(* Logix 5000 project; controller PLC_MCC1201_220AP1 vendor 1 type 14 code 164 rev 35.11; software revision 35.00; part 5 of 25 *)
(* tags used below, declared in another part *)
   B3 : DINT[102];
   B52 : DINT[100];
   GP_OB_InitializeMain : GP_OB_Initialize;
   HMI_Alarm_Reset : BOOL;   // HMI_Alarm_Reset
   HMI_MAN_CMD_WR : UDT_MAN_CMD_WR;
   HOST_DATA_REQ : ALIAS FOR N43[209].0;
   I : INT[128];
   LEHR_SPEED : ALIAS FOR N60[1];
   M202_M1_DR : AXIS_CIP_DRIVE;
   M203_M1_DR : AXIS_CIP_DRIVE;
   M203DROP : MAC_DROPCONV;
   M203DROP_HMR : MAC_DROPCONV_HMR;
   M204_M1_DR : AXIS_CIP_DRIVE;
   M2xx_CONVEYOR : MAC_CONVEYOR[20];
   M2xx_CONVEYOR_IN_MOTION : MAC_CONVEYOR_IN_MOTION[20];
   M2xx_CONVEYOR_OUT_MOTION : MAC_CONVEYOR_OUT_MOTION[20];
   MS_ACCUM : ALIAS FOR N70[1];
   N : ALIAS FOR N15[80];
   N43 : DINT[240];
   N54 : DINT[501];
   N70 : DINT[3];
   N80 : DINT[16];
   O : INT[128];
   REL_CAP_REQUEST : ALIAS FOR I[17].14;
   S : INT[128];
   Status : INT;   // INT tag to retrieve Status value through GSV created during conversion
   T4 : TIMER[100];
   T57 : TIMER[100];
   TMP_dDirection : DINT;
   TMP_rAcc : REAL;
   TMP_rDec : REAL;
   TMP_rSpeed : REAL;
   TMP_xAlwaysOFF : BOOL;
   TMP_xRun : BOOL;
   W_B3 : DINT[7];

   W_CONV_MSG_N7_0 : MESSAGE;   // IFE1_BTW_CNT
        .EN   // btw_enable
        MessageParameters(ServiceCode := 16#004c, LocalElement := W_N7[10], ...)
   W_CONV_MSG_N7_120 : MESSAGE;   // OFE1_CONTROL
        .EN   // BTW_OFE1_ENABLE
        MessageParameters(ServiceCode := 16#004c, LocalElement := W_N7[140], ...)
   W_CONV_MSG_N7_160 : MESSAGE;   // OFE1_BTR_CONTRO
        .EN   // OFE1_BTR_ENABLE
        MessageParameters(ServiceCode := 16#004b, LocalElement := W_N7[180], ...)
   W_CONV_MSG_N7_200 : MESSAGE;   // OFE2_CONTROL
        .EN   // OFE2_BTW_ENABLE
        MessageParameters(ServiceCode := 16#004c, LocalElement := W_N7[220], ...)
   W_CONV_MSG_N7_240 : MESSAGE;   // OFE2_BTR_CONTRO
        .EN   // OFE2_BTR_ENABLE
        MessageParameters(ServiceCode := 16#004b, LocalElement := W_N7[260], ...)
   W_CONV_MSG_N7_280 : MESSAGE;   // OFE3_CONTROL
        .EN   // OFE3_BTW_ENABLE
        MessageParameters(ServiceCode := 16#004c, LocalElement := W_N7[300], ...)
   W_CONV_MSG_N7_32 : MESSAGE;   // IFE1_BTR
        .EN   // BTR_IFE1_ENABLE
        MessageParameters(ServiceCode := 16#004b, LocalElement := W_N7[42], ...)
   W_CONV_MSG_N7_320 : MESSAGE;   // OFE3_BTR_CONTRL
        .EN   // OFE3_BTR_ENABLE
        MessageParameters(ServiceCode := 16#004b, LocalElement := W_N7[340], ...)
   W_CONV_MSG_N7_360 : MESSAGE;   // OFE4_CONTROL
        .EN   // OFE4_BTW_CONTRL
        MessageParameters(ServiceCode := 16#004c, LocalElement := W_N7[380], ...)
   W_CONV_MSG_N7_400 : MESSAGE;   // OFE4_BTR_CONTRL
        .EN   // OFE4_BTR_ENABLE
        MessageParameters(ServiceCode := 16#004b, LocalElement := W_N7[420], ...)
   W_CONV_MSG_N7_60 : MESSAGE;   // IFE2_CONTROL
        .EN   // IFE2_BTW_ENABLE
        MessageParameters(ServiceCode := 16#004c, LocalElement := W_N7[70], ...)
   W_CONV_MSG_N7_92 : MESSAGE;   // IFE2_BTR
        .EN   // BTR_IFE2_ENABLE
        MessageParameters(ServiceCode := 16#004b, LocalElement := W_N7[102], ...)
   W_CONV_PID_N7_440 : PID := (CTL := 1115722368, CT := 1, CA := 1, PE := 1, INI := 1, OLH := 1, DVPA := 1, PVHA := 1, SP := 2048.0, KP := 500.0, BIAS := 2973.0, MAXS := 4095.0, SO := 100.0, MAXO := 100.0, UPD := 1.0, PV := 4095.0, ERR := 2047.0, OUT := 100.0, MAXI := 4095.0, MAXTIE := 4095.0, DATA[1] := 1600.0, DATA[2] := 4095.0, DATA[3] := 2047.0, DATA[4] := 2048.0, DATA[5] := 0.024420025, DATA[6] := 1.0, DATA[7] := 16.0, DATA[8] := 500.0, DATA[11] := 500.0, DATA[16] := 0.024420025);   // Receiving Tank Level Control
   W_CONV_PID_N7_470 : PID := (CTL := 1082168192, CT := 1, PE := 1, INI := 1, OLH := 1, DVPA := 1, PVLA := 1, PVHA := 1, SP := 1845.0, KP := 150.0, KI := 300.0, BIAS := 2045.0, MAXS := 4095.0, SO := 100.0, MAXO := 100.0, UPD := 1.0, ERR := 1845.0, OUT := 100.0, MAXI := 4095.0, MAXTIE := 4095.0, DATA[3] := 1845.0, DATA[4] := 1845.0, DATA[5] := 0.024420025, DATA[6] := 1.0, DATA[7] := 16.0, DATA[8] := 150.0, DATA[9] := 300.0, DATA[11] := 150.0, DATA[12] := 0.008333334, DATA[16] := 0.024420025);   // Washer Water Pressure Cntrl Valve Position
   W_CONV_PID_N7_500 : PID := (CTL := 1082168192, CT := 1, PE := 1, INI := 1, OLH := 1, DVPA := 1, PVLA := 1, PVHA := 1, SP := 2050.0, KP := 250.0, BIAS := 2045.0, MAXS := 4095.0, SO := 100.0, MAXO := 100.0, UPD := 1.0, ERR := 2050.0, OUT := 100.0, MAXI := 4095.0, MAXTIE := 4095.0, DATA[3] := 2050.0, DATA[4] := 2050.0, DATA[5] := 0.024420025, DATA[6] := 1.0, DATA[7] := 16.0, DATA[8] := 250.0, DATA[11] := 250.0, DATA[16] := 0.024420025);   // Dryer Room Airflow (CB2) Fan Actuator Control
   W_CONV_PID_N7_530 : PID := (CTL := 8430720, PE := 1, INI := 1, OLL := 1, DVNA := 1, PVHA := 1, SP := 2073.0, KP := 100.0, KI := 300.0, BIAS := 2047.0, MAXS := 4095.0, MAXO := 100.0, UPD := 1.0, PV := 4095.0, ERR := -2022.0, MAXI := 4095.0, MAXTIE := 4095.0, DATA[1] := -1600.0, DATA[2] := 4095.0, DATA[3] := -2022.0, DATA[4] := 2073.0, DATA[5] := 0.024420025, DATA[6] := 1.0, DATA[7] := 16.0, DATA[8] := 100.0, DATA[9] := 300.0, DATA[11] := 100.0, DATA[12] := 0.0055555557, DATA[16] := 0.024420025);   // Blower CB1 Static Pressure Fan Actuator Control
   W_CONV_PID_N7_560 : PID := (CTL := 8430720, PE := 1, INI := 1, OLL := 1, DVNA := 1, PVHA := 1, SP := 1023.0, KP := 300.0, KI := 300.0, BIAS := 2047.0, MAXS := 4095.0, MAXO := 100.0, UPD := 1.0, PV := 1339.0, ERR := -316.0, MAXI := 4095.0, MAXTIE := 4095.0, DATA[1] := -523.1746, DATA[2] := 1339.0, DATA[3] := -316.0, DATA[4] := 1023.0, DATA[5] := 0.024420025, DATA[6] := 1.0, DATA[7] := 16.0, DATA[8] := 300.0, DATA[9] := 300.0, DATA[11] := 300.0, DATA[12] := 0.016666668, DATA[16] := 0.024420025);   // RO Heating Coil Temp. Control (HC1)
   W_CONV_PID_N7_590 : PID := (CTL := 1082167936, CT := 1, PE := 1, INI := 1, OLH := 1, DVPA := 1, PVHA := 1, SP := 2559.0, KP := 250.0, KI := 300.0, BIAS := 2047.0, MAXS := 4095.0, SO := 100.0, MAXO := 100.0, UPD := 1.0, PV := 525.0, ERR := 2034.0, OUT := 100.0, MAXI := 4095.0, MAXTIE := 4095.0, DATA[1] := -205.1282, DATA[2] := 525.0, DATA[3] := 2034.0, DATA[4] := 2559.0, DATA[5] := 0.024420025, DATA[6] := 1.0, DATA[7] := 16.0, DATA[8] := 250.0, DATA[9] := 300.0, DATA[11] := 250.0, DATA[12] := 0.013888889, DATA[16] := 0.024420025);   // Eclipse Heating Coil Temp. Control
   W_CONV_PID_N7_620 : PID := (CTL := 1082168192, CT := 1, PE := 1, INI := 1, OLH := 1, DVPA := 1, PVLA := 1, PVHA := 1, SP := 615.0, KP := 500.0, KI := 300.0, BIAS := 2047.0, MAXS := 4095.0, SO := 100.0, MAXO := 100.0, UPD := 1.0, ERR := 615.0, OUT := 100.0, MAXI := 4095.0, MAXTIE := 4095.0, DATA[3] := 615.0, DATA[4] := 615.0, DATA[5] := 0.024420025, DATA[6] := 1.0, DATA[7] := 16.0, DATA[8] := 500.0, DATA[9] := 300.0, DATA[11] := 500.0, DATA[12] := 0.027777778, DATA[16] := 0.024420025);   // Return Water Flow Control Valve Position
   W_CONV_PID_N7_650 : PID := (CTL := 41985152, CA := 1, PE := 1, INI := 1, OLL := 1, DVNA := 1, PVHA := 1, SP := 1971.0, KP := 400.0, KI := 100.0, BIAS := 2047.0, MAXS := 4095.0, MAXO := 100.0, UPD := 1.0, PV := 1713.0, ERR := -258.0, MAXI := 4095.0, MAXTIE := 4095.0, DATA[1] := 669.304, DATA[2] := 1713.0, DATA[3] := -258.0, DATA[4] := 1971.0, DATA[5] := 0.024420025, DATA[6] := 1.0, DATA[7] := 16.0, DATA[8] := 400.0, DATA[9] := 100.0, DATA[11] := 400.0, DATA[12] := 0.06666667, DATA[16] := 0.024420025);   // RO Unit Water Temperature Control
   W_CONV_PID_N7_680 : PID := (CTL := 1082167936, CT := 1, PE := 1, INI := 1, OLH := 1, DVPA := 1, PVHA := 1, SP := 2047.0, KP := 300.0, KI := 300.0, BIAS := 2047.0, MAXS := 4095.0, SO := 100.0, MAXO := 100.0, UPD := 1.0, PV := 439.0, ERR := 1608.0, OUT := 100.0, MAXI := 4095.0, MAXTIE := 4095.0, DATA[1] := -171.52626, DATA[2] := 439.0, DATA[3] := 1608.0, DATA[4] := 2047.0, DATA[5] := 0.024420025, DATA[6] := 1.0, DATA[7] := 16.0, DATA[8] := 300.0, DATA[9] := 300.0, DATA[11] := 300.0, DATA[12] := 0.016666668, DATA[16] := 0.024420025);   // Boiler Water Temperature Control
   W_CONV_PID_N7_710 : PID := (CTL := 1082167936, CT := 1, PE := 1, INI := 1, OLH := 1, DVPA := 1, PVHA := 1, SP := 2047.0, KP := 300.0, KI := 200.0, BIAS := 2047.0, MAXS := 4095.0, SO := 100.0, MAXO := 100.0, UPD := 1.0, PV := 1029.0, ERR := 1018.0, OUT := 100.0, MAXI := 4095.0, MAXTIE := 4095.0, DATA[1] := -402.0513, DATA[2] := 1029.0, DATA[3] := 1018.0, DATA[4] := 2047.0, DATA[5] := 0.024420025, DATA[6] := 1.0, DATA[7] := 16.0, DATA[8] := 300.0, DATA[9] := 200.0, DATA[11] := 300.0, DATA[12] := 0.025, DATA[16] := 0.024420025);   // Mixed Air Control Damper Positioning
   W_CONV_PID_N7_740 : PID := (CTL := 1082168192, CT := 1, PE := 1, INI := 1, OLH := 1, DVPA := 1, PVLA := 1, PVHA := 1, SP := 1024.0, KP := 300.0, KI := 300.0, BIAS := 2047.0, MAXS := 4095.0, SO := 100.0, MAXO := 100.0, UPD := 1.0, ERR := 1024.0, OUT := 100.0, MAXI := 4095.0, MAXTIE := 4095.0, DATA[3] := 1024.0, DATA[4] := 1024.0, DATA[5] := 0.024420025, DATA[6] := 1.0, DATA[7] := 16.0, DATA[8] := 300.0, DATA[9] := 300.0, DATA[11] := 300.0, DATA[12] := 0.016666668, DATA[16] := 0.024420025);   // Dryer Room Temperature Control
   W_CP1_ENABLE : ALIAS FOR W_B3[0].5;
   W_CP1A_START : ALIAS FOR W_O[10].5;
   W_CP1A_STATUS : ALIAS FOR W_I[8].7;
   W_CP1B_START : ALIAS FOR W_O[10].7;
   W_CP1B_STATUS : ALIAS FOR W_I[8].6;
   W_CP2A_START : ALIAS FOR W_O[10].9;
   W_CP2A_STAT : ALIAS FOR W_I[8].4;
   W_CP2B_START : ALIAS FOR W_O[10].11;
   W_CP2B_STAT : ALIAS FOR W_I[8].3;
   W_DRV_OUTPUT : ALIAS FOR W_N7[380];
   W_DRV_PID : ALIAS FOR W_N7[440];
   W_DRYER_AIR_FLOW : ALIAS FOR W_N7[108];
   W_DRYER_PID_OUT : ALIAS FOR W_N7[925];
   W_DRYER_TEMP_PID : ALIAS FOR W_N7[740];
   W_DRYER_TEMP_TMR : ALIAS FOR W_T4[16];
   W_EMER_STOP : ALIAS FOR W_I[8].13;
   W_EMER_STOP_LIGHT : ALIAS FOR W_O[10].10;
   W_F8 : REAL[1];
   W_FAN_CB1_TIMER : ALIAS FOR W_T4[4];
   W_FAN_CB2_TIMER : ALIAS FOR W_T4[5];
   W_FLOW_ENABLE : ALIAS FOR W_B3[0].9;
   W_HC1_SENSOR : ALIAS FOR W_N7[44];
   W_HEATING_AIR_ST : ALIAS FOR W_N7[107];
   W_HX1_BCD_OUT : ALIAS FOR W_N7[917];
   W_HX2_SENSOR : ALIAS FOR W_N7[47];
   W_I : INT[32] := ([8] := 2#0001_0000_0000_0110, [17] := 2#0000_0000_0101_0000);
        [16].8   // ?????????????? RO System Emergency Low Level Photoeye ??????????????
        [16].0   // Pump CP1A Drive Fault
        [16].1   // Pump CP1B Drive Fault
        [16].2   // RO Water Low Feed Pressure
        [16].3   // Reverse Osmosis Pump Motor Auxillary
        [16].4   // Eclipse On Selector at NSG Washer Panel (North)
        [16].5   // Eclipse Off Selector at NSG Washer Panel (North)
        [16].6   // Elipse On Selector at NSG Washer Panel (South)
        [16].7   // Eclipse Off Selector at NSG Washer Panel (South)
        [8].0   // Logical Shutdown Pushbutton
        [8].1   // Process Water Tank Low Level Limit Switch (Honeywell)
        [8].10   // APC Tank Fill Switch
        [8].11   // CB2 Blower Starter Auxillary
        [8].12   // CB1 Blower Starter Auxillary
        [8].13   // RO System Emergency Stop
        [8].14   // Pump CP1 Lead/Lag Switch
        [8].15   // Pump CP2 Lead/Lag Switch
        [8].2   // Process Water Tank High Limit
        [8].3   // CP2B Motor Starter Auxillary Status
        [8].4   // CP2A Motor Starter Auxillary Status
        [8].6   // CP1B Motor Auxillary Status
        [8].7   // CP1A Motor Auxillary Status
        [8].8   // PS1_Switch Pressure Switch
        [8].9   // Recieving Tank Level Switch (Cullet Tunnel)
        [8]   // WASHER INPUTS
        [16]   // WASHER INPUTS
   W_IFE1_BTW_CNT : ALIAS FOR W_N7[0];
   W_IFE1_BTW_DATA : ALIAS FOR W_N7[10];
   W_IFE2_BTR : ALIAS FOR W_N7[92];
   W_IFE2_CONTROL : ALIAS FOR W_N7[60];
   W_IFE2_DATA : ALIAS FOR W_N7[70];
   W_INT_FOR_BCD1 : ALIAS FOR W_N7[911];
   W_LEVEL_SENSOR : ALIAS FOR W_N7[109];
   W_LL_CP1 : ALIAS FOR W_I[8].14;
   W_LL_CP1A_T : ALIAS FOR W_T4[2];
   W_LL_CP1B_T : ALIAS FOR W_T4[3];
   W_LL_CP2 : ALIAS FOR W_I[8].15;
   W_LL_CP2A_T : ALIAS FOR W_T4[0];
   W_LL_CP2B_T : ALIAS FOR W_T4[1];
   W_LL_TIMER : ALIAS FOR W_T4[100];
   W_LOG_SHUTDOWN : ALIAS FOR W_I[8].0;
   W_MA_FAN_SENSOR : ALIAS FOR W_N7[50];
   W_MIX_AIR_PID : ALIAS FOR W_N7[710];
   W_N11 : DINT[10] := ([0] := 11, [1] := 15);
        [0].0   // Host Read Log Shutdown Latch Enabled
        [0].1   // Host Read Run Washer
        [0].2   // Host Read RO System Emergency Stop
        [0].3   // Host Read RO System Pump Motor Started
        [0].4   // Host Read APC Active
        [0].5   // Host Read Blowdown Valve Energized
        [0].6   // Host Read RO Water Pump Motor Auxillary
        [1].0   // Host Read Pump CP2A Motor Started
        [1].1   // Host Read Pump CP2B Motor Started
        [1].2   // Host Read Process Water Tank Low Limit Detected
        [1].3   // Host Read Process Water Tank High Limit Detected
        [1].4   // Host Read Receiving Level Warning
        [1].5   // Host Read RO Water Low Feed Pressure
        [2].0   // Host Read CP1 Enabled
        [2].1   // Host Read Pump CP1A Drive Started
        [2].2   // Host Read Pump CP1A Drive Fault
        [2].3   // Host Read Pump CP1B Drive Started
        [2].4   // Host Read Pump CP1B Drive Fault
        [2].5   // Host Read Spare Pump On Signal Detected
        [2].6   // Host Read Flow Enable
        [2].7   // Host Read PS1 Enabled
        [3].0   // Host Read Fan CB1 Started
        [3].1   // Host Read Fan CB2 Started
   W_N189 : DINT[40] := ([0] := 29);
   W_N7 : DINT[933] := ([0] := 25624, [1] := 3, [2] := 3, [3] := 7, [4] := 10, [12] := 256, [16] := 16533, [18] := 16533, [20] := 16533, [22] := 16533, [24] := 16533, [26] := 16533, [28] := 16533, [30] := 16533, [31] := 12, [32] := -4456, [33] := 12, [34] := 12, [35] := 7, [36] := 42, [42] := 2, [43] := 36, [46] := 4921, [47] := 1081, [49] := 5907, [50] := 4137, [52] := 4760, [53] := 1317, [60] := 25628, [61] := 3, [62] := 3, [63] := 7, [64] := 70, [72] := 256, [76] := 16533, [78] := 16533, [80] := 16533, [82] := 16533, [84] := 16533, [86] := 16533, [88] := 16533, [90] := 16533, [91] := 12, [92] := -4452, [93] := 12, [94] := 12, [95] := 7, [96] := 102, [102] := 2, [103] := 245, [104] := 10, [107] := 16533, [109] := 16533, [120] := -4608, [121] := 13, [122] := 13, [123] := 7, [124] := 140, [136] := 16533, [138] := 16533,
        [143] := 7, [146] := 16533, [148] := 16533, [150] := 16533, [152] := 16533, [153] := 7, [154] := 160, [160] := -4480, [161] := 5, [162] := 5, [163] := 7, [164] := 180, [176] := 256, [178] := 256, [181] := 4095, [182] := 4095, [183] := 7, [184] := 64, [196] := 16533, [198] := 16533, [200] := -4604, [201] := 13, [202] := 13, [203] := 7, [204] := 220, [210] := 2052, [211] := 5, [213] := 7, [214] := 220, [216] := 256, [218] := 256, [226] := 16533, [228] := 16533, [230] := 16533, [232] := 16533, [240] := -4476, [241] := 5, [242] := 5, [243] := 7, [244] := 260, [256] := 16533, [258] := 16533, [260] := 4095, [263] := 4095, [264] := 64, [270] := 2056, [271] := 5, [273] := 7, [274] := 280, [280] := -4600, [281] := 13, [282] := 13, [283] := 7, [284] := 300, [293] := 10, [300] := 16533, [303] := 16533, [306] := 16533, [308] := 16533, [310] := 16533,
        [312] := 16533, [313] := 10, [316] := 16533, [318] := 16533, [320] := -4472, [321] := 5, [322] := 5, [323] := 7, [324] := 340, [330] := 2060, [331] := 5, [333] := 7, [334] := 340, [340] := 4095, [341] := 4095, [342] := 4095, [344] := 64, [353] := 1, [360] := -4596, [361] := 13, [362] := 13, [363] := 7, [364] := 380, [386] := 16533, [388] := 16533, [390] := 16533, [392] := 16533, [400] := -4468, [401] := 5, [402] := 5, [403] := 7, [404] := 420, [420] := 4095, [424] := 64, [440] := 557, [442] := 2048, [443] := 500, [446] := 2973, [447] := 4095, [450] := 100, [451] := 100, [453] := 1, [454] := 4095, [455] := 2047, [456] := 100, [459] := 99, [460] := -1600, [461] := 2047, [462] := 2048, [463] := 1, [470] := -24055, [471] := 100, [472] := 1845, [473] := 150, [474] := 300, [476] := 2045, [477] := 4095, [481] := 100, [483] := 1, [485] := 1845,
        [486] := 100, [491] := 1845, [492] := 1845, [493] := 1, [500] := 545, [502] := 2050, [503] := 250, [506] := 2045, [507] := 4095, [511] := 100, [513] := 1, [515] := 2050, [516] := 100, [521] := 2050, [522] := 2050, [523] := 1, [530] := 1033, [531] := 100, [532] := 2073, [533] := 100, [534] := 300, [536] := 2047, [537] := 4095, [541] := 100, [543] := 1, [544] := 4095, [545] := -2022, [547] := -14321, [548] := 21912, [549] := -100, [550] := 1600, [551] := -2022, [552] := 2073, [553] := 1, [560] := 1065, [561] := 1, [562] := 1023, [563] := 300, [564] := 300, [566] := 2047, [567] := 4095, [570] := 100, [571] := 100, [573] := 1, [574] := 1339, [575] := -316, [577] := -13600, [578] := -21394, [579] := -33, [580] := 20288, [581] := -925, [582] := 1023, [583] := 7, [584] := 380, [590] := 553, [591] := 1, [592] := 2559, [593] := 250, [594] := 300, [596] := 2047,
        [597] := 4095, [601] := 100, [603] := 1, [604] := 522, [605] := 2037, [606] := 100, [609] := -13, [610] := 16768, [611] := 1478, [612] := 2559, [620] := 553, [621] := 1, [622] := 615, [623] := 500, [624] := 300, [626] := 2047, [627] := 4095, [631] := 100, [633] := 1, [635] := 615, [636] := 100, [641] := 615, [642] := 615, [650] := 1037, [652] := 1971, [653] := 400, [654] := 100, [656] := 2047, [657] := 4095, [660] := 75, [661] := 100, [663] := 1, [664] := 1737, [665] := -234, [667] := -13531, [668] := 1444, [669] := 42, [670] := 26688, [671] := 1, [672] := 1971, [680] := 553, [682] := 2047, [683] := 300, [684] := 300, [686] := 2047, [687] := 4095, [691] := 100, [693] := 1, [695] := 2047, [696] := 100, [697] := 19002, [698] := 23044, [701] := 2039, [702] := 2047, [710] := 553, [712] := 2047, [713] := 300, [714] := 200, [716] := 2047, [717] := 4095,
        [721] := 100, [723] := 1, [724] := 1033, [725] := 1014, [726] := 100, [727] := 19255, [728] := 32691, [729] := -26, [730] := -14400, [731] := 230, [732] := 2047, [740] := 553, [742] := 1024, [743] := 300, [744] := 300, [746] := 2047, [747] := 4095, [751] := 100, [753] := 1, [755] := 1024, [756] := 100, [761] := 1024, [762] := 1024, [900] := 4095, [908] := 4095, [910] := 1339, [912] := 525, [916] := 1713, [918] := 439, [920] := 1029, [923] := 4095, [926] := 4095, [931] := 4095);
        [106]   // PT-1_Pressure
        [107]   // Heating_Air_St
        [108]   // Dryer_Air_Flow
        [109]   // Receiving Tank Level Transmit Value
        [10]   // IFE1_BTW_DATA
        [110]   // Conduct_Sensor
        [111]   // Sheet_Temp
        [140]   // Analog Output for Heat Exchng Temperature Control Valve
        [141]   // Analog Output for Boiler Water Temp. Control Valve
        [142]   // Analog Output Calculated for Pressure Cntl Valve Position Manipulation
        [180]   // OFE1_BTR_DATA
        [220]   // Analog Output for Return Water Flow Cntl Valve Positioning
        [221]   // Analog Output for APC Tank Valve Position
        [222]   // Analog Output For RO Heating Coil Damper Position
        [223]   // Analog Output for Eclipse Heating Coil Damper Position
        [260]   // OFE2_BTR_DATA
        [300]   // Analog Output to RET Temp. Conrol Damper
        [301]   // Analog Output to Lehr Temp. Control Damper
        [302]   // Analog Output for Dryer Room Temp. Control Damper 5A
        [303]   // Analog Output for Dryer Room Temp. Control Damper 5B
        [340]   // OFE3_BTR_DATA
        [380]   // Analog Output for Drive Control
        [382]   // Analog Output for CB1 Vortex Damper Position
        [383]   // Analog Output for CB2 Vortex Damper Position
        [420]   // OFE4_BTR_DATA
        [440].13   // test-btw
        [44]   // HC1_SENSOR
        [47]   // HX2_SENSOR
        [48]   // TT3_Raw_BCD
        [49]   // TT6_HITEMP_AIR
        [50]   // Mixed Air Control Sensor
        [51]   // TT8_SENSOR
        [53]   // TT8_RAW_DATA
        [70]   // IFE2_DATA
        [900]   // Receiving Tank Level Transmit Analog Input Value
        [902]   // Washer Water Pressure Transducer Analog Input Value
        [903]   // PID_to_Output
        [904]   // Drying Air Flow Measuring Station Analog Input Value
        [905]   // Drying Air Flow Value Square Root
        [906]   // Drying Air Flow Velocity
        [907]   // Out_From_Pid
        [908]   // Blower CB1 Static Pressure Probe Analog Input Value
        [910]   // RO Heating Coil Temp. Transmitter Analog Input Value
        [911]   // INT_FOR_TCD1
        [912]   // Eclipse Heat Coil Temp. Transmitter Analog Input Value
        [913]   // PID_BCD_TCD2
        [914]   // Return Water Conductivity Transmitter Analog Input Value
        [916]   // RO Unit Water Temperature Conrol Sensor Analog Input Value
        [917]   // HX1_OUT_BCD
        [918]   // Boiler Water Backup Heating Analog Input Value
        [919]   // PID_INT_TO_TOD
        [920]   // Mixed Air Temperature Transmitter Analog Input Value
        [921]   // RET_PID_OUTPUT
        [922]   // Mixed Air Temperature Control Damper Output
        [923]   // Compute Output to TCD3
        [924]   // Dryer Air Temperature Transmitter Analog Input Value
        [925]   // DRYER_PID_OUT
        [926]   // Compute Output to TCD5B
        [927]   // Reversed_Dryer
        [928]   // Fan CB2 Initialize
        [929]   // Fan CB1 Initialize
        [931]   // APC Tank Valve Position for Open
        [932]   // APC Tank Valve Position for Close
   W_O : INT[32] := ([10] := 2#0010_1010_0000_0000);
        [0]   // 12 Bit Ana log Output
        [10].1   // Fan CB1 Start
        [10].10   // Emergency Stop Light
        [10].11   // Pump CP2B Motor Start
        [10].12   // Signal to Open Blowdown Valve
        [10].13   // RO System Pump Motor Start
        [10].3   // Fan CB2 Start
        [10].5   // Pump CP1A Motor Start
        [10].7   // Pump CP1B Motor Start
        [10].8   // Receiving Tank Overflowing Warning Beacon
        [10].9   // Pump CP2A Motor Start
        [10]   // WASHER OUTPUTS
   W_OFE1_BTR_CONTRO : ALIAS FOR W_N7[160];
   W_OFE1_BTR_DATA : ALIAS FOR W_N7[180];
   W_OFE1_CONTROL : ALIAS FOR W_N7[120];
   W_OFE2_BTR_CONTRO : ALIAS FOR W_N7[240];
   W_OFE2_BTR_DATA : ALIAS FOR W_N7[260];
   W_OFE2_CONTROL : ALIAS FOR W_N7[200];
   W_OFE3_BTR_CONTRL : ALIAS FOR W_N7[320];
   W_OFE3_BTR_DATA : ALIAS FOR W_N7[340];
   W_OFE3_CONTROL : ALIAS FOR W_N7[280];
   W_OFE4_BTR_CONTRL : ALIAS FOR W_N7[400];
   W_OFE4_BTR_DATA : ALIAS FOR W_N7[420];
   W_OFE4_CONTROL : ALIAS FOR W_N7[360];
   W_OUT_FROM_PID : ALIAS FOR W_N7[907];
   W_PID_BCD_TCD2 : ALIAS FOR W_N7[913];
   W_PID_INT_TO_TOD : ALIAS FOR W_N7[919];
   W_PID_TO_OUTPUT : ALIAS FOR W_N7[903];
   W_PS1_SWITCH : ALIAS FOR W_I[8].8;
   W_PS1_TIMER : ALIAS FOR W_T4[50];
   W_PWT_HIGH_LIMIT : ALIAS FOR W_I[8].2;
   W_PWT_LL_LATCH : ALIAS FOR W_B3[0].8;
   W_R6 : CONTROL[1];
   W_RECIEVING_LEVEL : ALIAS FOR W_I[8].9;
   W_RET_PID_OUTPUT : ALIAS FOR W_N7[921];
   W_REVERSED_DRYER : ALIAS FOR W_N7[927];
   W_RO_SIG_START : ALIAS FOR W_B3[6].4;
   W_RO_START : ALIAS FOR W_O[10].13;
   W_RUN_WASHER : ALIAS FOR W_B3[0].2;
   W_S : INT[128] := ([1] := 16#2082, [2] := 16#d202, [8] := 16#0007, [9] := 16#0015, [10] := 16#0002, [18] := 16#0002, [19] := 16#0007, [20] := 16#0011, [21] := 16#0016, [22] := 16#0025, [23] := 16#0025, [28] := 16#01f4, [57] := 16#64a0, [78] := 16#0002, [80] := 16#0002, [81] := 16#0005, [82] := 16#0015, [83] := 16#0005, [84] := 16#0002, [85] := 16#0009);
        [0].0   // Processor arithmetic carry flag
        [0].1   // Processor arithmetic underflow/ overflow flag
        [0].2   // Processor arithmetic zero flag
        [0].3   // Processor arithmetic sign flag
        [100]   // Program G maximum scan time
        [101]   // Main control program H file number
        [102]   // Program H scan time
        [103]   // Program H maximum scan time
        [104]   // Main control program I file number
        [105]   // Program I scan time
        [106]   // Program I maximum scan time
        [107]   // Main control program J file number
        [108]   // Program J scan time
        [109]   // Program J maximum scan time
        [10].0   // Battery is bad or missing
        [10].1   // DH+ active node table changed
        [10].10   // MCP not allowed
        [10].11   // PII word number isn't in local rack
        [10].12   // User PII routine overlap
        [10].13   // No command block exists to get PII
        [10].14   // Arithmetic overflow occurred
        [10].15   // SFC lingering action overlap
        [10].2   // STI overlap
        [10].3   // EEPROM trans- ferred
        [10].4   // Edits prevent SFC continuing
        [10].5   // Invalid I/O status file
        [10].6   // Memory cartridge battery low
        [10].7   // No more command blocks exist
        [10].9   // No MCP was configured to run
        [110]   // Main control program K file number
        [111]   // Program K scan time
        [112]   // Program K maximum scan time
        [113]   // Main control program L file number
        [114]   // Program L scan time
        [115]   // Program L maximum scan time
        [116]   // Main control program M file number
        [117]   // Program M scan time
        [118]   // Program M maximum scan time
        [119]   // Main control program N file number
        [11].0   // Bad program file
        [11].1   // Bad address in ladder program
        [11].10   // Hardware Error
        [11].11   // MCP file does not exist or is not ladder
        [11].12   // PII file does not exist or is not ladder
        [11].13   // STI file does not exist or is not ladder
        [11].14   // Fault file does not exist or is not ladder
        [11].15   // Non ladder file
        [11].2   // Programmer error
        [11].3   // SFC Fault
        [11].4   // Program assembly error
        [11].5   // Powerup protection fault
        [11].6   // Error not defined
        [11].7   // User generated fault
        [11].8   // Watchdog timer fault
        [11].9   // Bad system config- uration
        [120]   // Program N scan time
        [121]   // Program N maximum scan time
        [122]   // Main control program O file number
        [123]   // Program O scan time
        [124]   // Program O maximum scan time
        [125]   // Main control program P file number
        [126]   // Program P scan time
        [127]   // Program P maximum scan time
        [12]   // Fault Code
        [13]   // Program file where fault occurred
        [14]   // Rung number where fault occurred
        [16]   // I/O status file
        [17].0   // Queue full between local and remote I/O
        [17].1   // Queue full servicing channel 1A
        [17].2   // Queue full servicing channel 1B
        [17].3   // Queue full servicing channel 2A
        [17].4   // Queue full servicing channel 2B
        [17].5   // No modem on serial port
        [17].6   // Remote I/O is greater than image size
        [17].8   // ASCII instruct- ion error
        [17].9   // Duplicate node address
        [18]   // Real time clock YEAR
        [19]   // Real time clock MONTH
        [1].0   // Bad RAM CHECKSUM at power up
        [1].1   // PLC-5 in RUN mode
        [1].10   // EEPROM success- fully Burned
        [1].11   // Perform- ing online program- ming
        [1].12   // Processor is in DEBUG mode
        [1].13   // User program CHECKSUM done
        [1].14   // Last scan of ladder or SFC step
        [1].15   // First scan of ladder or SFC step
        [1].2   // PLC-5 in TEST mode
        [1].3   // PLC-5 in PROG mode
        [1].4   // PLC-5 is burning an EEPROM
        [1].5   // Download- ing in progress
        [1].6   // Test edits enabled
        [1].7   // Mode switch in REMOTE
        [1].8   // Forces enabled
        [1].9   // Forces present
        [20]   // Real time clock DAY
        [21]   // Real time clock HOUR
        [22]   // Real time clock MINUTE
        [23]   // Real time clock SECOND
        [24]   // Indexed Addressing Offset
        [25]   // Adapter Image File
        [26].0   // SFC Restart/ Continue
        [26].1   // Start-up protect- ion after power loss
        [26].2   // Local rack is 1 if set or 0 if bit = 0
        [26].3   // Complement Rack Mode
        [27].0   // Rack 0 Inhibit
        [27].1   // Rack 1 Inhibit
        [27].10   // Rack 2 Reset
        [27].11   // Rack 3 Reset
        [27].12   // Rack 4 Reset
        [27].13   // Rack 5 Reset
        [27].14   // Rack 6 Reset
        [27].15   // Rack 7 Reset
        [27].2   // Rack 2 Inhibit
        [27].3   // Rack 3 Inhibit
        [27].4   // Rack 4 Inhibit
        [27].5   // Rack 5 Inhibit
        [27].6   // Rack 6 Inhibit
        [27].7   // Rack 7 Inhibit
        [27].8   // Rack 0 Reset
        [27].9   // Rack 1 Reset
        [28]   // Watchdog Timer Setpoint
        [29]   // Fault routine file number
        [30]   // STI setpoint (interval)
        [31]   // STI file number
        [32].0   // Rack 10 Faulted
        [32].1   // Rack 11 Faulted
        [32].10   // Block Xfer queue to rack 12 is full
        [32].11   // Block Xfer queue to rack 13 is full
        [32].12   // Block Xfer queue to rack 14 is full
        [32].13   // Block Xfer queue to rack 15 is full
        [32].14   // Block Xfer queue to rack 16 is full
        [32].15   // Block Xfer queue to rack 17 is full
        [32].2   // Rack 12 Faulted
        [32].3   // Rack 13 Faulted
        [32].4   // Rack 14 Faulted
        [32].5   // Rack 15 Faulted
        [32].6   // Rack 16 Faulted
        [32].7   // Rack 17 Faulted
        [32].8   // Block Xfer queue to rack 10 is full
        [32].9   // Block Xfer queue to rack 11 is full
        [33].0   // Rack 10 Inhibit
        [33].1   // Rack 11 Inhibit
        [33].10   // Rack 12 Reset
        [33].11   // Rack 13 Reset
        [33].12   // Rack 14 Reset
        [33].13   // Rack 15 Reset
        [33].14   // Rack 16 Reset
        [33].15   // Rack 17 Reset
        [33].2   // Rack 12 Inhibit
        [33].3   // Rack 13 Inhibit
        [33].4   // Rack 14 Inhibit
        [33].5   // Rack 15 Inhibit
        [33].6   // Rack 16 Inhibit
        [33].7   // Rack 17 Inhibit
        [33].8   // Rack 10 Reset
        [33].9   // Rack 11 Reset
        [34].0   // Rack 20 Faulted
        [34].1   // Rack 21 Faulted
        [34].10   // Block Xfer queue to rack 22 is full
        [34].11   // Block Xfer queue to rack 23 is full
        [34].12   // Block Xfer queue to rack 24 is full
        [34].13   // Block Xfer queue to rack 25 is full
        [34].14   // Block Xfer queue to rack 26 is full
        [34].15   // Block Xfer queue to rack 27 is full
        [34].2   // Rack 22 Faulted
        [34].3   // Rack 23 Faulted
        [34].4   // Rack 24 Faulted
        [34].5   // Rack 25 Faulted
        [34].6   // Rack 26 Faulted
        [34].7   // Rack 27 Faulted
        [34].8   // Block Xfer queue to rack 20 is full
        [34].9   // Block Xfer queue to rack 21 is full
        [35].0   // Rack 20 Inhibit
        [35].1   // Rack 21 Inhibit
        [35].10   // Rack 22 Reset
        [35].11   // Rack 23 Reset
        [35].12   // Rack 24 Reset
        [35].13   // Rack 25 Reset
        [35].14   // Rack 26 Reset
        [35].15   // Rack 27 Reset
        [35].2   // Rack 22 Inhibit
        [35].3   // Rack 23 Inhibit
        [35].4   // Rack 24 Inhibit
        [35].5   // Rack 25 Inhibit
        [35].6   // Rack 26 Inhibit
        [35].7   // Rack 27 Inhibit
        [35].8   // Rack 20 Reset
        [35].9   // Rack 21 Reset
        [46]   // PII file number
        [47]   // PII module group to examine
        [48]   // PII bit mask
        [48].0   // PII Module Bit 1=Monitor 0=Ignore
        [49]   // PII compare value
        [49].0   // PII Bit 1=false to true, 0= true to false
        [50]   // PII down count
        [51]   // PII return mask
        [52]   // PII accum- ulator
        [53]   // STI last scan time
        [54]   // STI max scan time
        [55]   // PII last scan time
        [56]   // PII max scan time
        [79].0   // Main control program A disable bit
        [79].1   // Main control program B disable bit
        [79].10   // Main control program K disable bit
        [79].11   // Main control program L disable bit
        [79].12   // Main control program M disable bit
        [79].13   // Main control program N disable bit
        [79].14   // Main control program O disable bit
        [79].15   // Main control program P disable bit
        [79].2   // Main control program C disable bit
        [79].3   // Main control program D disable bit
        [79].4   // Main control program E disable bit
        [79].5   // Main control program F disable bit
        [79].6   // Main control program G disable bit
        [79].7   // Main control program H disable bit
        [79].8   // Main control program I disable bit
        [79].9   // Main control program J disable bit
        [7].0   // Rack 0 Faulted
        [7].1   // Rack 1 Faulted
        [7].10   // Block Xfer queue to rack 2 is full
        [7].11   // Block Xfer queue to rack 3 is full
        [7].12   // Block Xfer queue to rack 4 is full
        [7].13   // Block Xfer queue to rack 5 is full
        [7].14   // Block Xfer queue to rack 6 is full
        [7].15   // Block Xfer queue to rack 7 is full
        [7].2   // Rack 2 Faulted
        [7].3   // Rack 3 Faulted
        [7].4   // Rack 4 Faulted
        [7].5   // Rack 5 Faulted
        [7].6   // Rack 6 Faulted
        [7].7   // Rack 7 Faulted
        [7].8   // Block Xfer queue to rack 0 is full
        [7].9   // Block Xfer queue to rack 1 is full
        [80]   // Main control program A file number
        [81]   // Program A scan time
        [82]   // Program A maximum scan time
        [83]   // Main control program B file number
        [84]   // Program B scan time
        [85]   // Program B maximum scan time
        [86]   // Main control program C file number
        [87]   // Program C scan time
        [88]   // Program C maximum scan time
        [89]   // Main control program D file number
        [8]   // Last program scan time ladder & SFC
        [90]   // Program D scan time
        [91]   // Program D maximum scan time
        [92]   // Main control program E file number
        [93]   // Program E scan time
        [94]   // Program E maximum scan time
        [95]   // Main control program F file number
        [96]   // Program F scan time
        [97]   // Program F maximum scan time
        [98]   // Main control program G file number
        [99]   // Program G scan time
        [9]   // Maximum program scan time ladder & SFC
   W_SHEET_TEMP : ALIAS FOR W_N7[111];
   W_SHUTDOWN_LATCH : ALIAS FOR W_B3[0].1;
   W_SIG_CP1A_START : ALIAS FOR W_B3[0].6;
   W_SIG_CP1B_START : ALIAS FOR W_B3[0].7;
   W_SIG_CP2A_START : ALIAS FOR W_B3[0].3;
   W_SIG_CP2B_START : ALIAS FOR W_B3[0].4;
   W_T4 : TIMER[101] := ([0].PRE := 20000, [1].PRE := 20000, [1].ACC := 20000, [1].EN := 1, [1].DN := 1, [2].PRE := 20000, [3].PRE := 20000, [4].PRE := 30000, [5].PRE := 20000, [6].PRE := 100, [6].ACC := 20, [6].EN := 1, [6].TT := 1, [7].PRE := 100, [7].ACC := 20, [7].EN := 1, [7].TT := 1, [8].PRE := 100, [8].ACC := 20, [8].EN := 1, [8].TT := 1, [9].PRE := 100, [9].ACC := 20, [9].EN := 1, [9].TT := 1, [10].PRE := 100, [10].ACC := 20, [10].EN := 1, [10].TT := 1, [11].PRE := 100, [11].ACC := 20, [11].EN := 1, [11].TT := 1, [12].PRE := 100, [12].ACC := 20, [12].EN := 1, [12].TT := 1, [13].PRE := 100, [13].ACC := 20, [13].EN := 1, [13].TT := 1, [14].PRE := 100, [14].ACC := 20, [14].EN := 1, [14].TT := 1, [15].PRE := 100, [15].ACC := 20, [15].EN := 1, [15].TT := 1, [16].PRE := 100, [16].ACC := 20, [16].EN := 1, [16].TT := 1, [17].PRE := 3600000, [17].ACC := 879250, [17].EN := 1, [17].TT := 1, [18].PRE := 15000, [20].PRE := 300000, [24].PRE := 30000,
        [25].PRE := 14400000, [25].ACC := 4479270, [25].EN := 1, [25].TT := 1, [26].PRE := 14400000, [50].PRE := 60000, [99].PRE := 300000, [100].PRE := 300000, [100].ACC := 300000, [100].EN := 1, [100].DN := 1);
        [0]   // CP2A Pump Motor Start-up Failure Timer
        [0].DN   // LL_CP2A_T
        [100]   // Process Water Tank Low Limit Timer
        [10]   // RO Water Heating Coil (HC1) Timer
        [11]   // Eclipse Heating Coil (HC2) Timer
        [12]   // Return Water Conductivity Timer
        [13]   // RO Unit Water Heat Exchanger (HX1) Timer
        [14]   // Boiler Water Backup Heating Timer
        [15]   // Blower Timer
        [16]   // Dryer Room Temperature Timer
        [17]   // Blowdown Valve Cycle Timer
        [18]   // Blowdown Valve Active Duration Timer
        [18].TT   // Blowdown_ON
        [1]   // CP2B Pump Motor Start-up Failure Timer
        [1].DN   // LL_CP2B_T
        [20]   // APC Tank Fill Cycle Timer
        [20].DN   // APC Tank Fill Cycle Done
        [25]   // Process Water Timer to Switch Active Pump 4 Hours On
        [26]   // Process Water Timer to Switch Active Pump 4 Hours Off
        [2]   // CP1A Motor Start-up Failure Timer
        [2].DN   // CP1_LL_TIMER
        [3]   // CP1B Motor Start-up Failure Timer
        [3].DN   // CP1B_LL_TIMER
        [4]   // Delay to Start Fan CB1
        [50]   // Pressure Switch 1 Timer
        [5]   // Delay to Start Fan CB2
        [6]   // Receiving Tank Level (CP1 Pumps) PID Timer
        [7]   // Pressure Control Valve Timer
        [8]   // Dryer Room Airflow PID Timer
        [99]   // Timer to delay the Emergency low level alarm horn
        [9]   // Blower CB1 Static Pressure Timer
   W_TCD1_OUTPUT : ALIAS FOR W_N7[222];
   W_TCD1_PID : ALIAS FOR W_N7[560];
   W_TCD2_OUTPUT : ALIAS FOR W_N7[223];
   W_TCD2_PID : ALIAS FOR W_N7[590];
   W_TCD3_OUTPUT : ALIAS FOR W_N7[300];
   W_TCD3_PID_OUTPUT : ALIAS FOR W_N7[922];
   W_TCD4_OUTPUT : ALIAS FOR W_N7[301];
   W_TCD5A_OUTPUT : ALIAS FOR W_N7[302];
   W_TMP_xAlwaysOFF : BOOL; {access Read Only}
   W_TT3_RAW_BCD : ALIAS FOR W_N7[48];
   W_TT6_HITEMP_AIR : ALIAS FOR W_N7[49];
   W_TT8_INPUT : ALIAS FOR W_N7[912];
   W_TT8_RAW_DATA : ALIAS FOR W_N7[53];
   W_TT8_SENSOR : ALIAS FOR W_N7[51];
   W_WARNING_LIGHT : ALIAS FOR W_O[10].8;
   WASH_AK1_CON : ALIAS FOR N54[203].4;
   WASH_AK1_CR : ALIAS FOR N54[207].4;
   WASH_AK1_RET : ALIAS FOR N54[203].3;
   WASH_AK1_SV : ALIAS FOR O[36].2;
   WASH_AK1LO_CVG : ALIAS FOR N54[206].4;
   WASH_AK1UP_CVG : ALIAS FOR N54[205].4;
   WASH_AK2_CON : ALIAS FOR N54[203].6;
   WASH_AK2_CR : ALIAS FOR N54[207].5;
   WASH_AK2_RET : ALIAS FOR N54[203].5;
   WASH_AK2_SV : ALIAS FOR O[36].0;
   WASH_AK2LO_CVG : ALIAS FOR N54[206].5;
   WASH_AK2UP_CVG : ALIAS FOR N54[205].5;
   WASH_ARK_AUTO : ALIAS FOR N54[203].1;
   WASH_ARK_MANLMP : ALIAS FOR N54[203].9;
   WASH_ARK_MANUAL : ALIAS FOR N54[203].2;
   WASH_BR1_AUTO : ALIAS FOR N54[200].1;
   WASH_BR1_CR : ALIAS FOR N54[207].1;
   WASH_BR1_CRT : ALIAS FOR T57[1];
   WASH_BR1_MANLMP : ALIAS FOR N54[200].9;
   WASH_BR1_MANUAL : ALIAS FOR N54[200].2;
   WASH_BR1_MOFF : ALIAS FOR N54[200].10;
   WASH_BR1_OFF : ALIAS FOR N54[200].4;
   WASH_BR1_ON : ALIAS FOR N54[200].3;
   WASH_BR1_SPY : ALIAS FOR N54[205].6;
   WASH_BR1_SV : ALIAS FOR O[36].12;
   WASH_BR1LO_CON : ALIAS FOR N54[200].8;
   WASH_BR1LO_CVG : ALIAS FOR N54[206].1;
   WASH_BR1LO_RET : ALIAS FOR N54[200].7;
   WASH_BR1UP_CON : ALIAS FOR N54[200].6;
   WASH_BR1UP_CVG : ALIAS FOR N54[205].1;
   WASH_BR1UP_RET : ALIAS FOR N54[200].5;
   WASH_BR1UP_SV : ALIAS FOR O[36].14;
   WASH_BR2_CR : ALIAS FOR N54[207].2;
   WASH_BR2_CRT : ALIAS FOR T57[2];
   WASH_BR2_SPY : ALIAS FOR N54[205].7;
   WASH_CR_ACK : ALIAS FOR N54[207].0;
   WASH_CR_RESET : ALIAS FOR N54[207].7;
   WASH_MSTR_SPY : ALIAS FOR N54[205].9;
   WASH_SPG_AUTO : ALIAS FOR N54[202].1;
   WASH_SPG_CR : ALIAS FOR N54[207].3;
   WASH_SPG_MANLMP : ALIAS FOR N54[202].9;
   WASH_SPG_MANUAL : ALIAS FOR N54[202].2;
   WASH_SPG_MOFF : ALIAS FOR N54[202].10;
   WASH_SPG_OFF : ALIAS FOR N54[202].4;
   WASH_SPG_ON : ALIAS FOR N54[202].3;
   WASH_SPG_SPY : ALIAS FOR N54[205].8;
   WASH_SPGLO_CON : ALIAS FOR N54[202].8;
   WASH_SPGLO_CVG : ALIAS FOR N54[206].3;
   WASH_SPGLO_RET : ALIAS FOR N54[202].7;
   WASH_SPGLO_SV : ALIAS FOR O[36].4;
   WASH_SPGUP_CON : ALIAS FOR N54[202].6;
   WASH_SPGUP_CVG : ALIAS FOR N54[205].3;
   WASH_SPGUP_RET : ALIAS FOR N54[202].5;
   WASH_SPGUP_SV : ALIAS FOR O[36].6;
   WASH_SPY3_TMR : ALIAS FOR T57[6];
   WASH_SPY_AUTO : ALIAS FOR N54[204].1;
   WASH_SPY_MANLMP : ALIAS FOR N54[204].9;
   WASH_SPY_MANUAL : ALIAS FOR N54[204].2;
   WASH_SPY_OFF : ALIAS FOR N54[204].4;
   WASH_SPY_ON : ALIAS FOR N54[204].3;
   WASH_SPYLO_CON : ALIAS FOR N54[204].8;
   WASH_SPYLO_RET : ALIAS FOR N54[204].7;
   WASH_SPYUP_CON : ALIAS FOR N54[204].6;
   WASH_SPYUP_RET : ALIAS FOR N54[204].5;
   WATER1_ON : ALIAS FOR O[47].7;
   WATER2_ON : ALIAS FOR O[47].8;
   WATER3_CR : ALIAS FOR N54[207].6;
   WATER3_ON : ALIAS FOR O[47].9;